(* Logix 5000 project; controller NWGG 1756-L72 rev 35.12; software revision 35.00; part 19 of 19 *)
(* tags used below, declared in another part *)
   Auto_Start_Treatment : BOOL;
   B_Offset : REAL;
   Bins_Rqd : BOOL;
   Blow_Out_Time : DINT;
   Blow_Out_Time_Remaining : REAL;
   Clean_Bin_Gates_Opened : BOOL;
   DeltaX : REAL;
   DeltaY : REAL;
   IDX : DINT;
   Loadout_Bin : udt_Loadout_Bin[29];
   Loadout_K_Valve : udt_Loadout_K_Valve[2];
   Loop_Idx : DINT;
   Manual_Blow_Out : BOOL;
   Manual_Open_Calibration_Valves : BOOL;
   Manually_Start_Treater : BOOL;
   Pause_Treatment : BOOL;
   Point1 : DINT;
   Point2 : DINT;
   Rate_Mult : REAL;
   Slope : REAL;
   Test1 : BOOL;
   tmr_Auto_Start : TIMER;
   tmr_Blow_Out : TIMER;
   Treat_Batch_Status : DINT;
   Treater_Calibration : BOOL;
   Treater_Loadout : udt_Treater_Loadout;
   Treatment_Running : BOOL;
   X1 : REAL;
   X2 : REAL;
   Y1 : REAL;
   Y2 : REAL;
   _700_TREAT : ALIAS FOR I7.3;
   test : BOOL;
   Treater_Remote_In : DINT;
   Treater_Remote_Out : DINT;
(* SeedLoadoutMain, continued *)

ROUTINE Treat_Bin_Gate_Ready   (* ladder *)
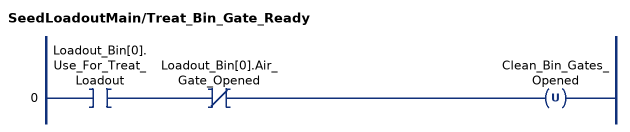
   0: XIC(Loadout_Bin[0].Use_For_Treat_Loadout)XIO(Loadout_Bin[0].Air_Gate_Opened)OTU(Clean_Bin_Gates_Opened);
END_ROUTINE

ROUTINE Treat_Bin_Rqd   (* ladder *)
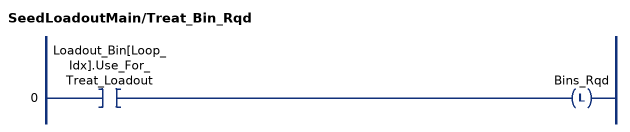
   0: XIC(Loadout_Bin[Loop_Idx].Use_For_Treat_Loadout)OTL(Bins_Rqd);
END_ROUTINE

ROUTINE Treaters   (* ladder *)
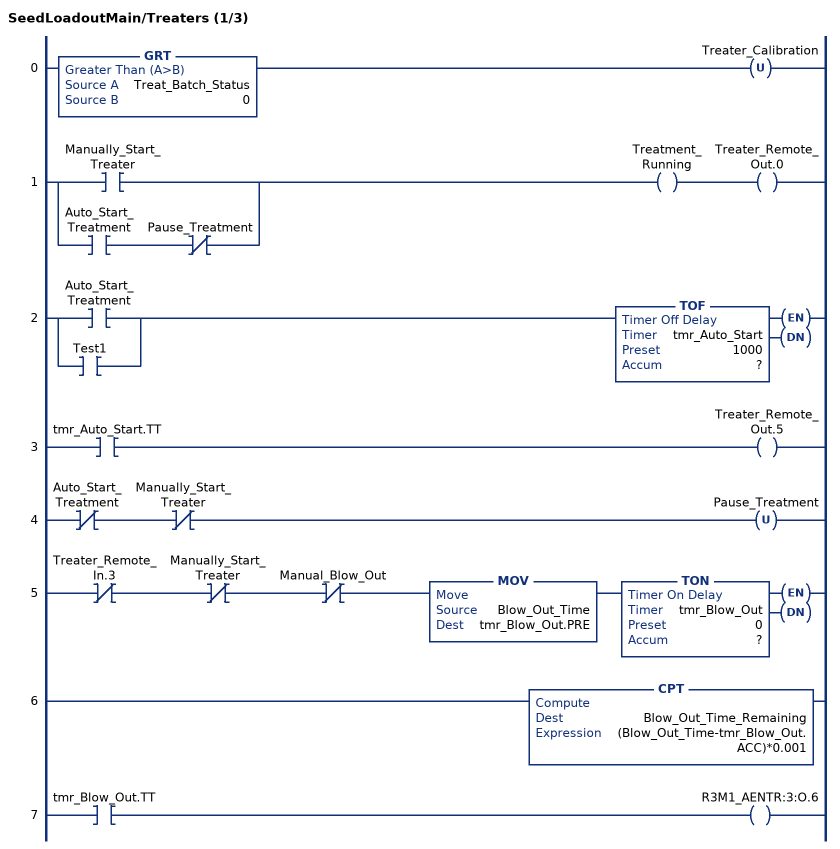
   0: GRT(Treat_Batch_Status,0)OTU(Treater_Calibration);
   1: [XIC(Manually_Start_Treater) ,XIC(Auto_Start_Treatment) XIO(Pause_Treatment) ]OTE(Treatment_Running)OTE(Treater_Remote_Out.0);
   2: [XIC(Auto_Start_Treatment) ,XIC(Test1) ]TOF(tmr_Auto_Start,?,?);
   3: XIC(tmr_Auto_Start.TT)OTE(Treater_Remote_Out.5);
   4: XIO(Auto_Start_Treatment)XIO(Manually_Start_Treater)OTU(Pause_Treatment);
   5: XIO(Treater_Remote_In.3)XIO(Manually_Start_Treater)XIO(Manual_Blow_Out)MOV(Blow_Out_Time,tmr_Blow_Out.PRE)TON(tmr_Blow_Out,?,?);
   6: CPT(Blow_Out_Time_Remaining,(Blow_Out_Time-tmr_Blow_Out.ACC)*0.001);
   7: XIC(tmr_Blow_Out.TT)OTE(R3M1_AENTR:3:O.6);
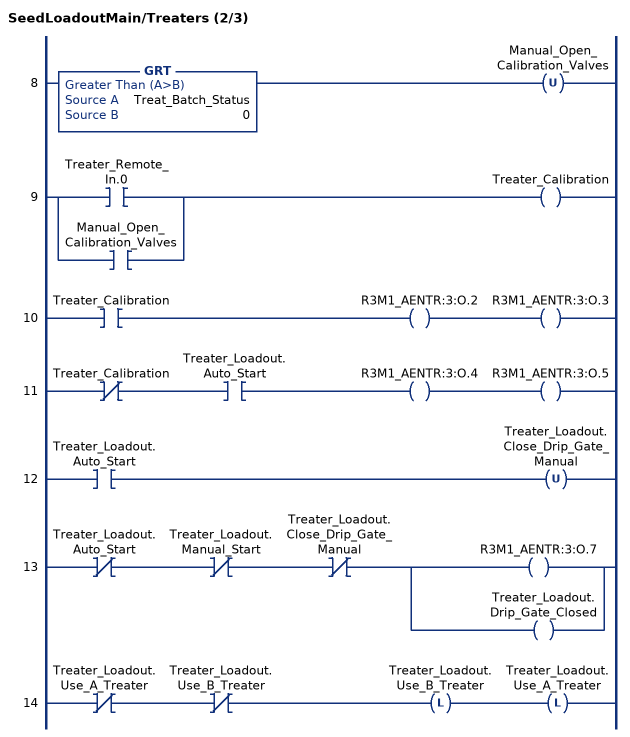
   8: GRT(Treat_Batch_Status,0)OTU(Manual_Open_Calibration_Valves);
   9: [XIC(Treater_Remote_In.0) ,XIC(Manual_Open_Calibration_Valves) ]OTE(Treater_Calibration);
   10: XIC(Treater_Calibration)OTE(R3M1_AENTR:3:O.2)OTE(R3M1_AENTR:3:O.3);
   11: XIO(Treater_Calibration)XIC(Treater_Loadout.Auto_Start)OTE(R3M1_AENTR:3:O.4)OTE(R3M1_AENTR:3:O.5);
   12: XIC(Treater_Loadout.Auto_Start)OTU(Treater_Loadout.Close_Drip_Gate_Manual);
   13: XIO(Treater_Loadout.Auto_Start)XIO(Treater_Loadout.Manual_Start)XIO(Treater_Loadout.Close_Drip_Gate_Manual)[OTE(R3M1_AENTR:3:O.7) ,OTE(Treater_Loadout.Drip_Gate_Closed) ];
   14: XIO(Treater_Loadout.Use_A_Treater)XIO(Treater_Loadout.Use_B_Treater)OTL(Treater_Loadout.Use_B_Treater)OTL(Treater_Loadout.Use_A_Treater);
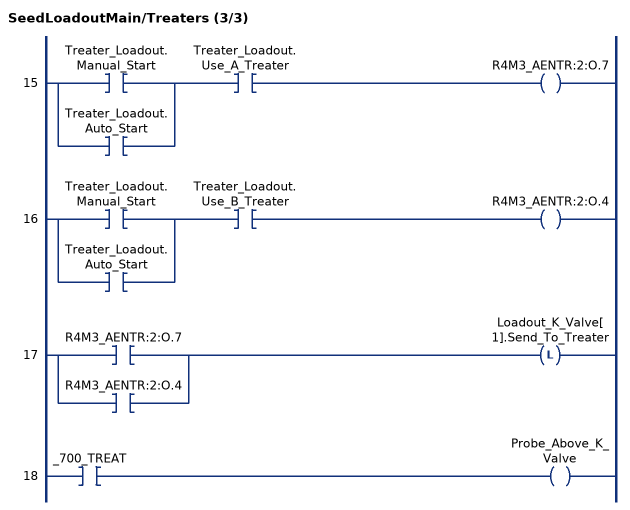
   15: [XIC(Treater_Loadout.Manual_Start) ,XIC(Treater_Loadout.Auto_Start) ]XIC(Treater_Loadout.Use_A_Treater)OTE(R4M3_AENTR:2:O.7);
   16: [XIC(Treater_Loadout.Manual_Start) ,XIC(Treater_Loadout.Auto_Start) ]XIC(Treater_Loadout.Use_B_Treater)OTE(R4M3_AENTR:2:O.4);
   17: [XIC(R4M3_AENTR:2:O.7) ,XIC(R4M3_AENTR:2:O.4) ]OTL(Loadout_K_Valve[1].Send_To_Treater);
   18: XIC(_700_TREAT)OTE(Probe_Above_K_Valve);
END_ROUTINE

ROUTINE Update_Andco_Cal_Points   (* ladder *)
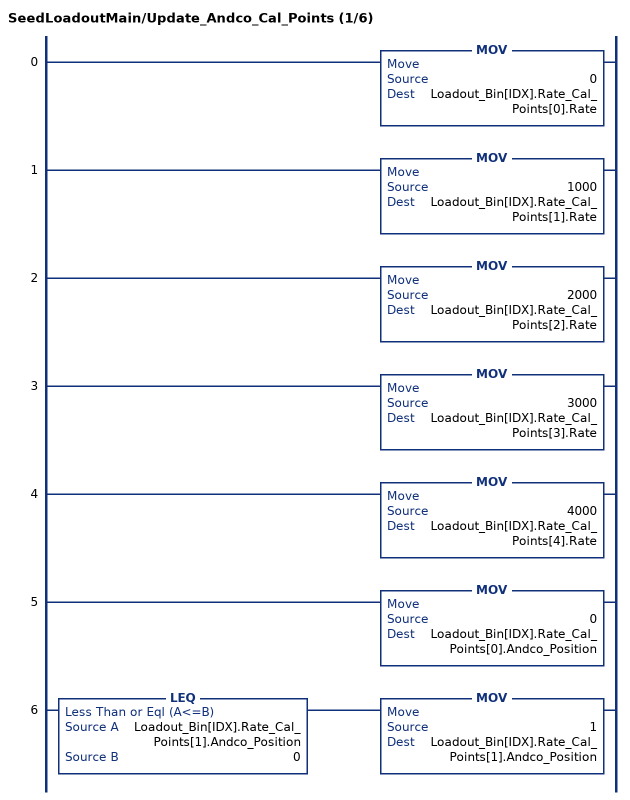
   0: MOV(0,Loadout_Bin[IDX].Rate_Cal_Points[0].Rate);
   1: MOV(1000,Loadout_Bin[IDX].Rate_Cal_Points[1].Rate);
   2: MOV(2000,Loadout_Bin[IDX].Rate_Cal_Points[2].Rate);
   3: MOV(3000,Loadout_Bin[IDX].Rate_Cal_Points[3].Rate);
   4: MOV(4000,Loadout_Bin[IDX].Rate_Cal_Points[4].Rate);
   5: MOV(0,Loadout_Bin[IDX].Rate_Cal_Points[0].Andco_Position);
   6: LEQ(Loadout_Bin[IDX].Rate_Cal_Points[1].Andco_Position,0)MOV(1,Loadout_Bin[IDX].Rate_Cal_Points[1].Andco_Position);
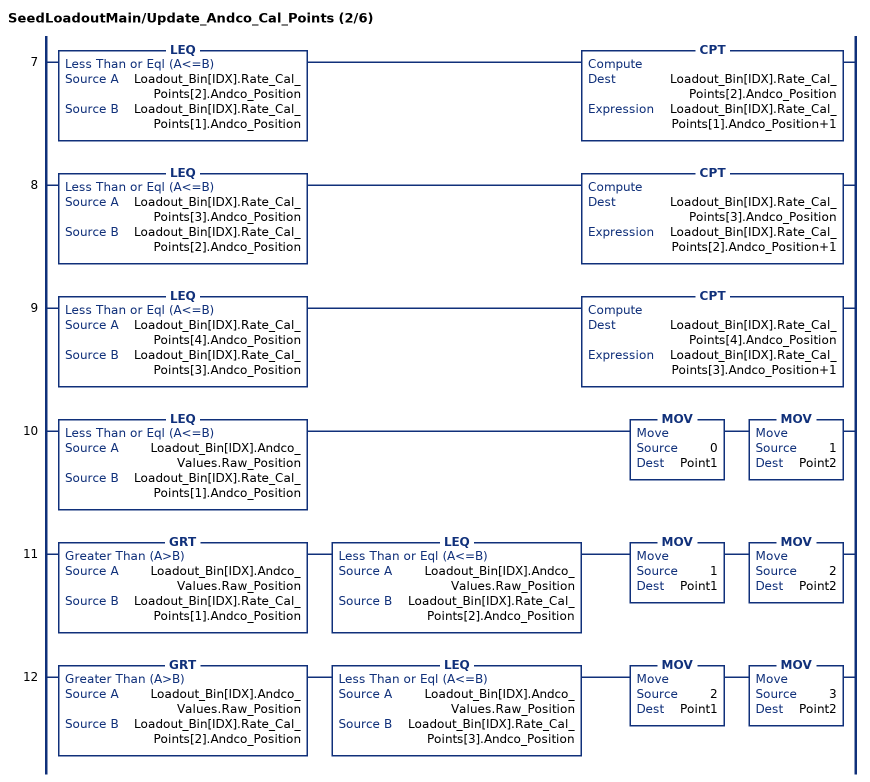
   7: LEQ(Loadout_Bin[IDX].Rate_Cal_Points[2].Andco_Position,Loadout_Bin[IDX].Rate_Cal_Points[1].Andco_Position)CPT(Loadout_Bin[IDX].Rate_Cal_Points[2].Andco_Position,Loadout_Bin[IDX].Rate_Cal_Points[1].Andco_Position+1);
   8: LEQ(Loadout_Bin[IDX].Rate_Cal_Points[3].Andco_Position,Loadout_Bin[IDX].Rate_Cal_Points[2].Andco_Position)CPT(Loadout_Bin[IDX].Rate_Cal_Points[3].Andco_Position,Loadout_Bin[IDX].Rate_Cal_Points[2].Andco_Position+1);
   9: LEQ(Loadout_Bin[IDX].Rate_Cal_Points[4].Andco_Position,Loadout_Bin[IDX].Rate_Cal_Points[3].Andco_Position)CPT(Loadout_Bin[IDX].Rate_Cal_Points[4].Andco_Position,Loadout_Bin[IDX].Rate_Cal_Points[3].Andco_Position+1);
   10: LEQ(Loadout_Bin[IDX].Andco_Values.Raw_Position,Loadout_Bin[IDX].Rate_Cal_Points[1].Andco_Position)MOV(0,Point1)MOV(1,Point2);
   11: GRT(Loadout_Bin[IDX].Andco_Values.Raw_Position,Loadout_Bin[IDX].Rate_Cal_Points[1].Andco_Position)LEQ(Loadout_Bin[IDX].Andco_Values.Raw_Position,Loadout_Bin[IDX].Rate_Cal_Points[2].Andco_Position)MOV(1,Point1)MOV(2,Point2);
   12: GRT(Loadout_Bin[IDX].Andco_Values.Raw_Position,Loadout_Bin[IDX].Rate_Cal_Points[2].Andco_Position)LEQ(Loadout_Bin[IDX].Andco_Values.Raw_Position,Loadout_Bin[IDX].Rate_Cal_Points[3].Andco_Position)MOV(2,Point1)MOV(3,Point2);
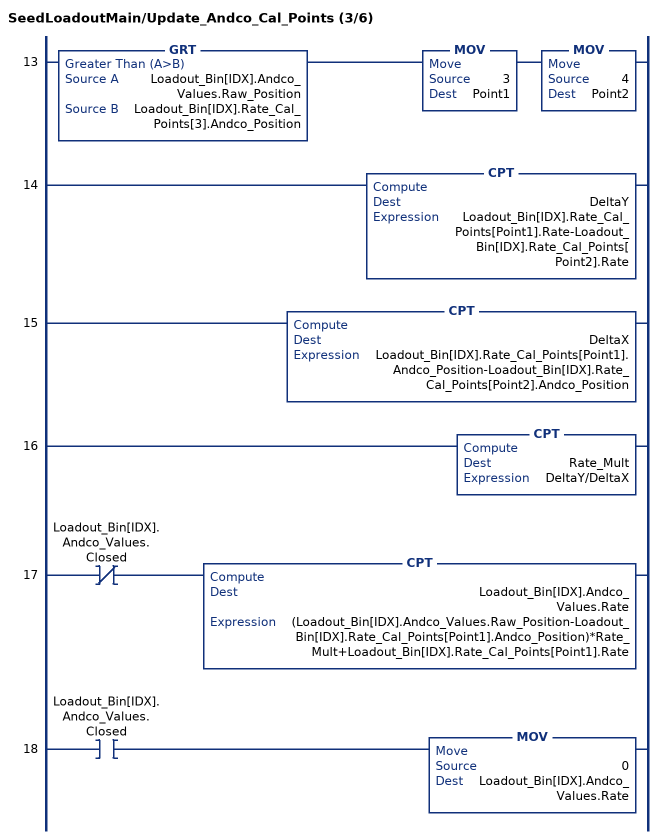
   13: GRT(Loadout_Bin[IDX].Andco_Values.Raw_Position,Loadout_Bin[IDX].Rate_Cal_Points[3].Andco_Position)MOV(3,Point1)MOV(4,Point2);
   14: CPT(DeltaY,Loadout_Bin[IDX].Rate_Cal_Points[Point1].Rate-Loadout_Bin[IDX].Rate_Cal_Points[Point2].Rate);
   15: CPT(DeltaX,Loadout_Bin[IDX].Rate_Cal_Points[Point1].Andco_Position-Loadout_Bin[IDX].Rate_Cal_Points[Point2].Andco_Position);
   16: CPT(Rate_Mult,DeltaY/DeltaX);
   17: XIO(Loadout_Bin[IDX].Andco_Values.Closed)CPT(Loadout_Bin[IDX].Andco_Values.Rate,(Loadout_Bin[IDX].Andco_Values.Raw_Position-Loadout_Bin[IDX].Rate_Cal_Points[Point1].Andco_Position)*Rate_Mult+Loadout_Bin[IDX].Rate_Cal_Points[Point1].Rate);
   18: XIC(Loadout_Bin[IDX].Andco_Values.Closed)MOV(0,Loadout_Bin[IDX].Andco_Values.Rate);
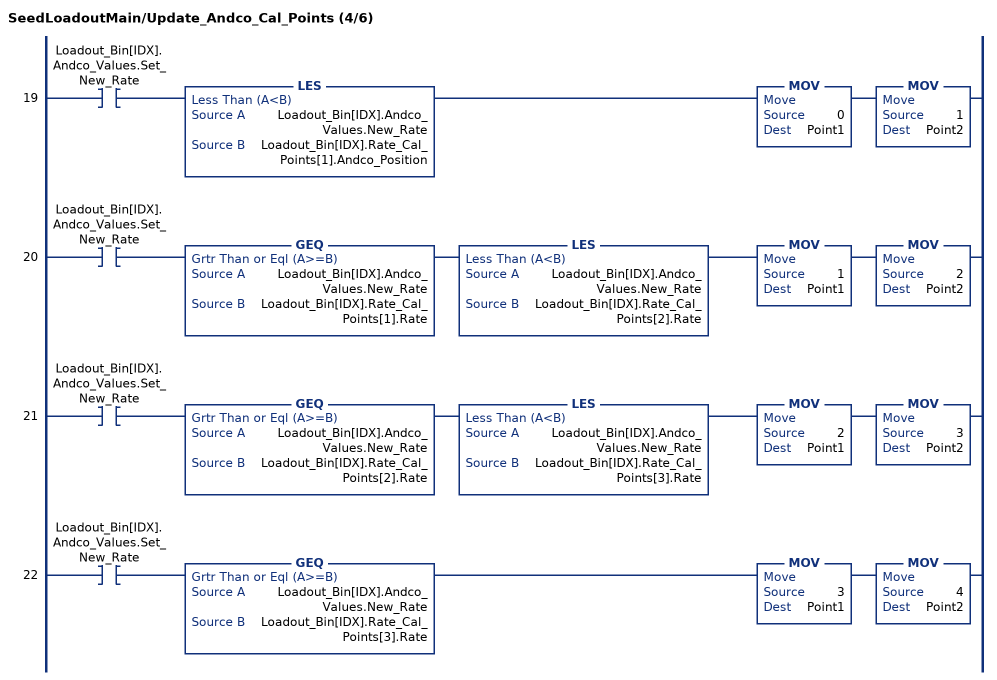
   19: XIC(Loadout_Bin[IDX].Andco_Values.Set_New_Rate)LES(Loadout_Bin[IDX].Andco_Values.New_Rate,Loadout_Bin[IDX].Rate_Cal_Points[1].Andco_Position)MOV(0,Point1)MOV(1,Point2);
   20: XIC(Loadout_Bin[IDX].Andco_Values.Set_New_Rate)GEQ(Loadout_Bin[IDX].Andco_Values.New_Rate,Loadout_Bin[IDX].Rate_Cal_Points[1].Rate)LES(Loadout_Bin[IDX].Andco_Values.New_Rate,Loadout_Bin[IDX].Rate_Cal_Points[2].Rate)MOV(1,Point1)MOV(2,Point2);
   21: XIC(Loadout_Bin[IDX].Andco_Values.Set_New_Rate)GEQ(Loadout_Bin[IDX].Andco_Values.New_Rate,Loadout_Bin[IDX].Rate_Cal_Points[2].Rate)LES(Loadout_Bin[IDX].Andco_Values.New_Rate,Loadout_Bin[IDX].Rate_Cal_Points[3].Rate)MOV(2,Point1)MOV(3,Point2);
   22: XIC(Loadout_Bin[IDX].Andco_Values.Set_New_Rate)GEQ(Loadout_Bin[IDX].Andco_Values.New_Rate,Loadout_Bin[IDX].Rate_Cal_Points[3].Rate)MOV(3,Point1)MOV(4,Point2);
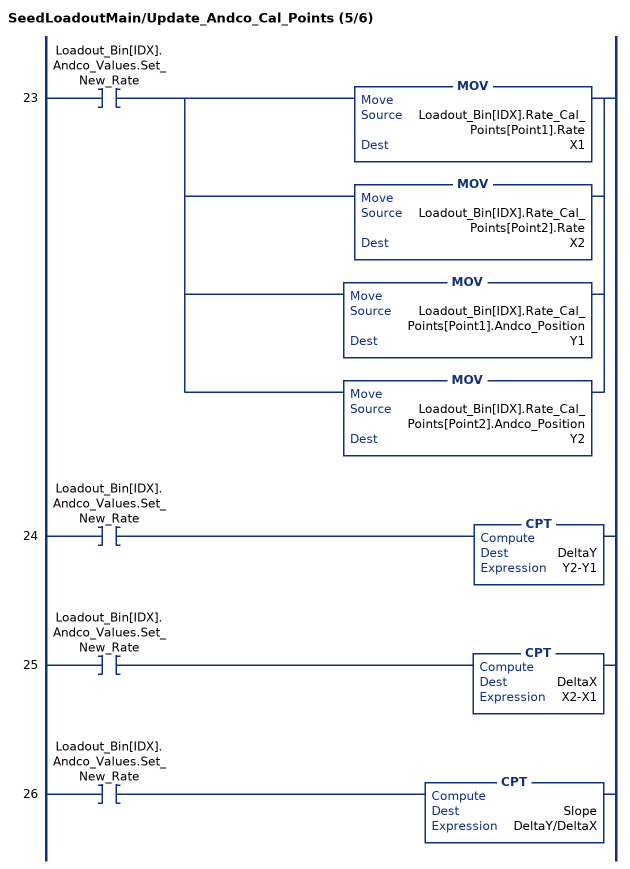
   23: XIC(Loadout_Bin[IDX].Andco_Values.Set_New_Rate)[MOV(Loadout_Bin[IDX].Rate_Cal_Points[Point1].Rate,X1) ,MOV(Loadout_Bin[IDX].Rate_Cal_Points[Point2].Rate,X2) ,MOV(Loadout_Bin[IDX].Rate_Cal_Points[Point1].Andco_Position,Y1) ,MOV(Loadout_Bin[IDX].Rate_Cal_Points[Point2].Andco_Position,Y2) ];
   24: XIC(Loadout_Bin[IDX].Andco_Values.Set_New_Rate)CPT(DeltaY,Y2-Y1);
   25: XIC(Loadout_Bin[IDX].Andco_Values.Set_New_Rate)CPT(DeltaX,X2-X1);
   26: XIC(Loadout_Bin[IDX].Andco_Values.Set_New_Rate)CPT(Slope,DeltaY/DeltaX);
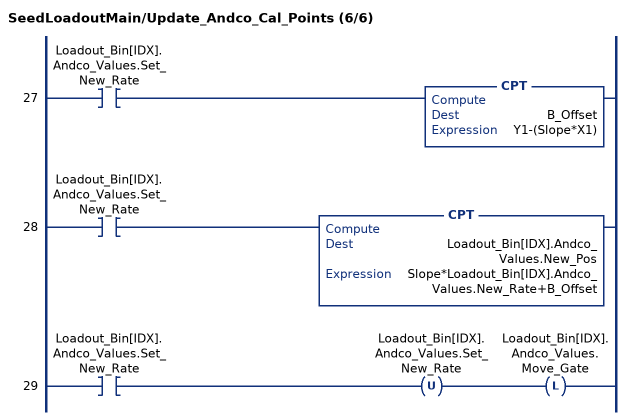
   27: XIC(Loadout_Bin[IDX].Andco_Values.Set_New_Rate)CPT(B_Offset,Y1-(Slope*X1));
   28: XIC(Loadout_Bin[IDX].Andco_Values.Set_New_Rate)CPT(Loadout_Bin[IDX].Andco_Values.New_Pos,Slope*Loadout_Bin[IDX].Andco_Values.New_Rate+B_Offset);
   29: XIC(Loadout_Bin[IDX].Andco_Values.Set_New_Rate)OTU(Loadout_Bin[IDX].Andco_Values.Set_New_Rate)OTL(Loadout_Bin[IDX].Andco_Values.Move_Gate);
END_ROUTINE
END_PROGRAM

PROGRAM Test   (* main routine Test *)
VAR
   Active : TIMER;
END_VAR

ROUTINE Test   (* ladder *)
END_ROUTINE
END_PROGRAM

PROGRAM Treating_NotUsed   (* main routine MainRoutine *)
VAR
   Probe_Above_K_Valve : BOOL;
END_VAR

ROUTINE MainRoutine   (* ladder *)
END_ROUTINE
END_PROGRAM

PROGRAM UpdateConfig
VAR
   BinIndex : DINT;
END_VAR
END_PROGRAM
